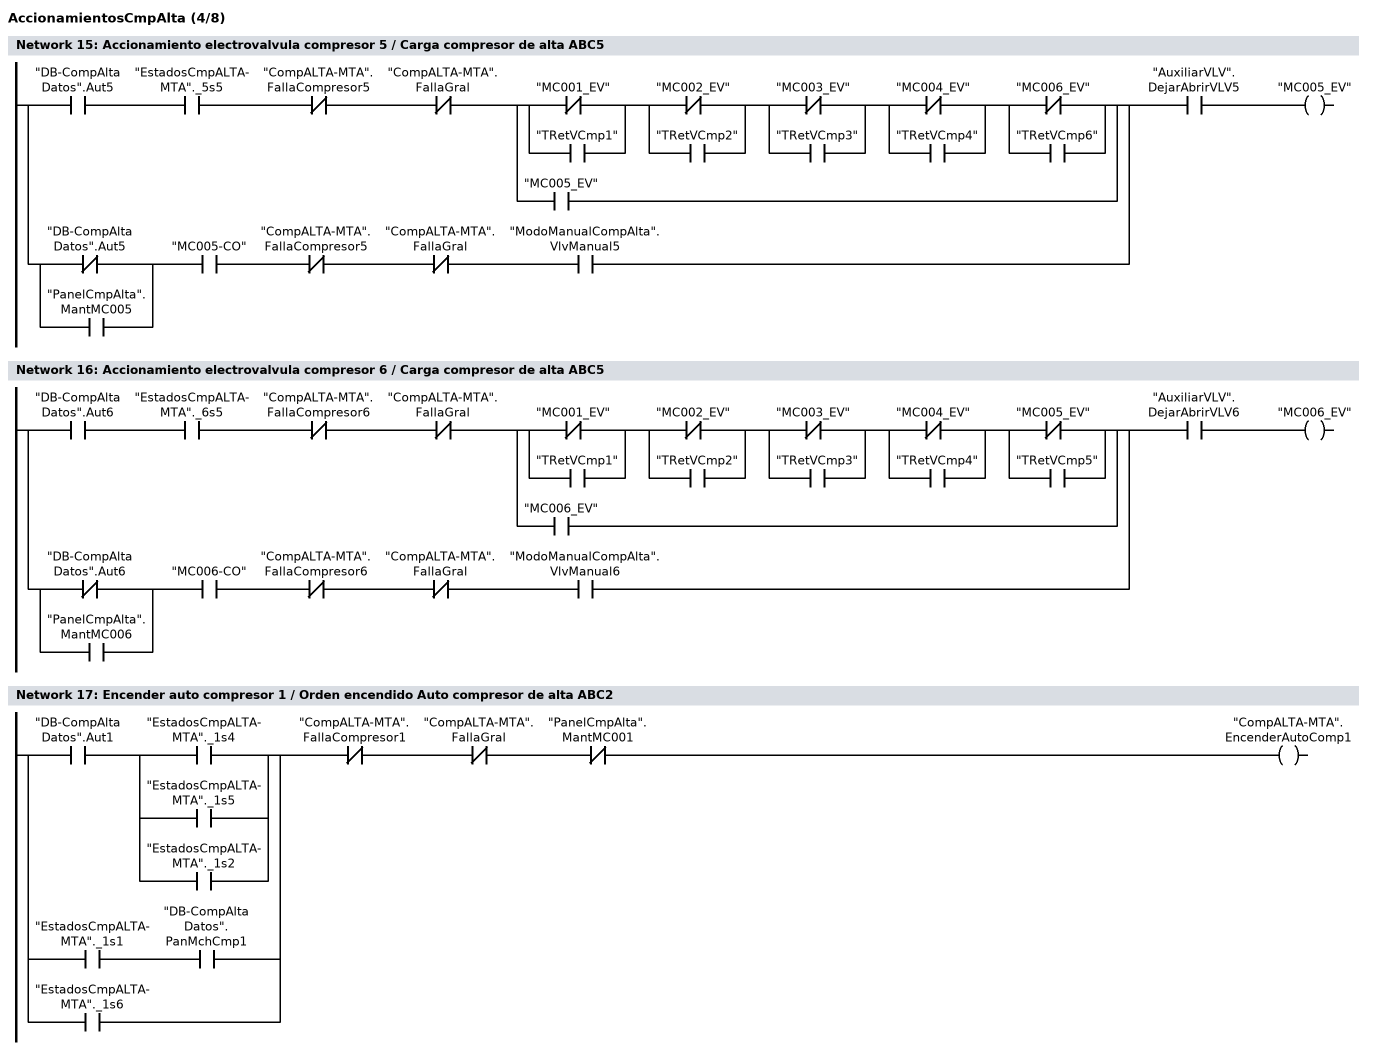
   RUNG wire#powerrail
      Contact( "DB-CompAltaDatos".Aut5 )
      Contact( "EstadosCmpALTA-MTA"._5s5 )
      I_Contact( "CompALTA-MTA".FallaCompresor5 )
      I_Contact( "CompALTA-MTA".FallaGral )
      wire#w1
      I_Contact( "MC001_EV" )
      wire#w2
      I_Contact( "MC002_EV" )
      wire#w3
      I_Contact( "MC003_EV" )
      wire#w4
      I_Contact( "MC004_EV" )
      wire#w5
      I_Contact( "MC006_EV" )
      wire#w6
      Contact( "AuxiliarVLV".DejarAbrirVLV5 )
      Coil( "MC005_EV" )
   END_RUNG
   RUNG wire#w1
      Contact( "TRetVCmp1" )
   END_RUNG wire#w2
   RUNG wire#w2
      Contact( "TRetVCmp2" )
   END_RUNG wire#w3
   RUNG wire#w3
      Contact( "TRetVCmp3" )
   END_RUNG wire#w4
   RUNG wire#w4
      Contact( "TRetVCmp4" )
   END_RUNG wire#w5
   RUNG wire#w5
      Contact( "TRetVCmp6" )
   END_RUNG wire#w6
   RUNG wire#w1
      Contact( "MC005_EV" )
   END_RUNG wire#w6
   RUNG wire#powerrail
      I_Contact( "DB-CompAltaDatos".Aut5 )
      wire#w7
      Contact( "MC005-CO" )
      I_Contact( "CompALTA-MTA".FallaCompresor5 )
      I_Contact( "CompALTA-MTA".FallaGral )
      Contact( "ModoManualCompAlta".VlvManual5 )
   END_RUNG wire#w6
   RUNG wire#powerrail
      Contact( "PanelCmpAlta".MantMC005 )
   END_RUNG wire#w7
   // the same network as SCL:
   "MC005_EV" := (("DB-CompAltaDatos".Aut5 AND "EstadosCmpALTA-MTA"._5s5 AND NOT "CompALTA-MTA".FallaCompresor5 AND NOT "CompALTA-MTA".FallaGral AND (((NOT "MC001_EV" OR "TRetVCmp1") AND (NOT "MC002_EV" OR "TRetVCmp2") AND (NOT "MC003_EV" OR "TRetVCmp3") AND (NOT "MC004_EV" OR "TRetVCmp4") AND (NOT "MC006_EV" OR "TRetVCmp6")) OR "MC005_EV")) OR ((NOT "DB-CompAltaDatos".Aut5 OR "PanelCmpAlta".MantMC005) AND "MC005-CO" AND NOT "CompALTA-MTA".FallaCompresor5 AND NOT "CompALTA-MTA".FallaGral AND "ModoManualCompAlta".VlvManual5)) AND "AuxiliarVLV".DejarAbrirVLV5;
END_REGION

REGION Network 16: Accionamiento electrovalvula compresor 6 / Carga compresor de alta ABC5
   RUNG wire#powerrail
      Contact( "DB-CompAltaDatos".Aut6 )
      Contact( "EstadosCmpALTA-MTA"._6s5 )
      I_Contact( "CompALTA-MTA".FallaCompresor6 )
      I_Contact( "CompALTA-MTA".FallaGral )
      wire#w1
      I_Contact( "MC001_EV" )
      wire#w2
      I_Contact( "MC002_EV" )
      wire#w3
      I_Contact( "MC003_EV" )
      wire#w4
      I_Contact( "MC004_EV" )
      wire#w5
      I_Contact( "MC005_EV" )
      wire#w6
      Contact( "AuxiliarVLV".DejarAbrirVLV6 )
      Coil( "MC006_EV" )
   END_RUNG
   RUNG wire#w1
      Contact( "TRetVCmp1" )
   END_RUNG wire#w2
   RUNG wire#w2
      Contact( "TRetVCmp2" )
   END_RUNG wire#w3
   RUNG wire#w3
      Contact( "TRetVCmp3" )
   END_RUNG wire#w4
   RUNG wire#w4
      Contact( "TRetVCmp4" )
   END_RUNG wire#w5
   RUNG wire#w5
      Contact( "TRetVCmp5" )
   END_RUNG wire#w6
   RUNG wire#w1
      Contact( "MC006_EV" )
   END_RUNG wire#w6
   RUNG wire#powerrail
      I_Contact( "DB-CompAltaDatos".Aut6 )
      wire#w7
      Contact( "MC006-CO" )
      I_Contact( "CompALTA-MTA".FallaCompresor6 )
      I_Contact( "CompALTA-MTA".FallaGral )
      Contact( "ModoManualCompAlta".VlvManual6 )
   END_RUNG wire#w6
   RUNG wire#powerrail
      Contact( "PanelCmpAlta".MantMC006 )
   END_RUNG wire#w7
   // the same network as SCL:
   "MC006_EV" := (("DB-CompAltaDatos".Aut6 AND "EstadosCmpALTA-MTA"._6s5 AND NOT "CompALTA-MTA".FallaCompresor6 AND NOT "CompALTA-MTA".FallaGral AND (((NOT "MC001_EV" OR "TRetVCmp1") AND (NOT "MC002_EV" OR "TRetVCmp2") AND (NOT "MC003_EV" OR "TRetVCmp3") AND (NOT "MC004_EV" OR "TRetVCmp4") AND (NOT "MC005_EV" OR "TRetVCmp5")) OR "MC006_EV")) OR ((NOT "DB-CompAltaDatos".Aut6 OR "PanelCmpAlta".MantMC006) AND "MC006-CO" AND NOT "CompALTA-MTA".FallaCompresor6 AND NOT "CompALTA-MTA".FallaGral AND "ModoManualCompAlta".VlvManual6)) AND "AuxiliarVLV".DejarAbrirVLV6;
END_REGION

REGION Network 17: Encender auto compresor 1 / Orden encendido Auto compresor de alta ABC2
   RUNG wire#powerrail
      Contact( "DB-CompAltaDatos".Aut1 )
      wire#w1
      Contact( "EstadosCmpALTA-MTA"._1s4 )
      wire#w2
      I_Contact( "CompALTA-MTA".FallaCompresor1 )
      I_Contact( "CompALTA-MTA".FallaGral )
      I_Contact( "PanelCmpAlta".MantMC001 )
      Coil( "CompALTA-MTA".EncenderAutoComp1 )
   END_RUNG
   RUNG wire#w1
      Contact( "EstadosCmpALTA-MTA"._1s5 )
   END_RUNG wire#w2
   RUNG wire#w1
      Contact( "EstadosCmpALTA-MTA"._1s2 )
   END_RUNG wire#w2
   RUNG wire#powerrail
      Contact( "EstadosCmpALTA-MTA"._1s1 )
      Contact( "DB-CompAltaDatos".PanMchCmp1 )
   END_RUNG wire#w2
   RUNG wire#powerrail
      Contact( "EstadosCmpALTA-MTA"._1s6 )
   END_RUNG wire#w2
   // the same network as SCL:
   "CompALTA-MTA".EncenderAutoComp1 := (("DB-CompAltaDatos".Aut1 AND ("EstadosCmpALTA-MTA"._1s4 OR "EstadosCmpALTA-MTA"._1s5 OR "EstadosCmpALTA-MTA"._1s2)) OR ("EstadosCmpALTA-MTA"._1s1 AND "DB-CompAltaDatos".PanMchCmp1) OR "EstadosCmpALTA-MTA"._1s6) AND NOT "CompALTA-MTA".FallaCompresor1 AND NOT "CompALTA-MTA".FallaGral AND NOT "PanelCmpAlta".MantMC001;
END_REGION

REGION Network 18: Encender auto compresor 2 / Orden encendido Auto compresor de alta ABC3
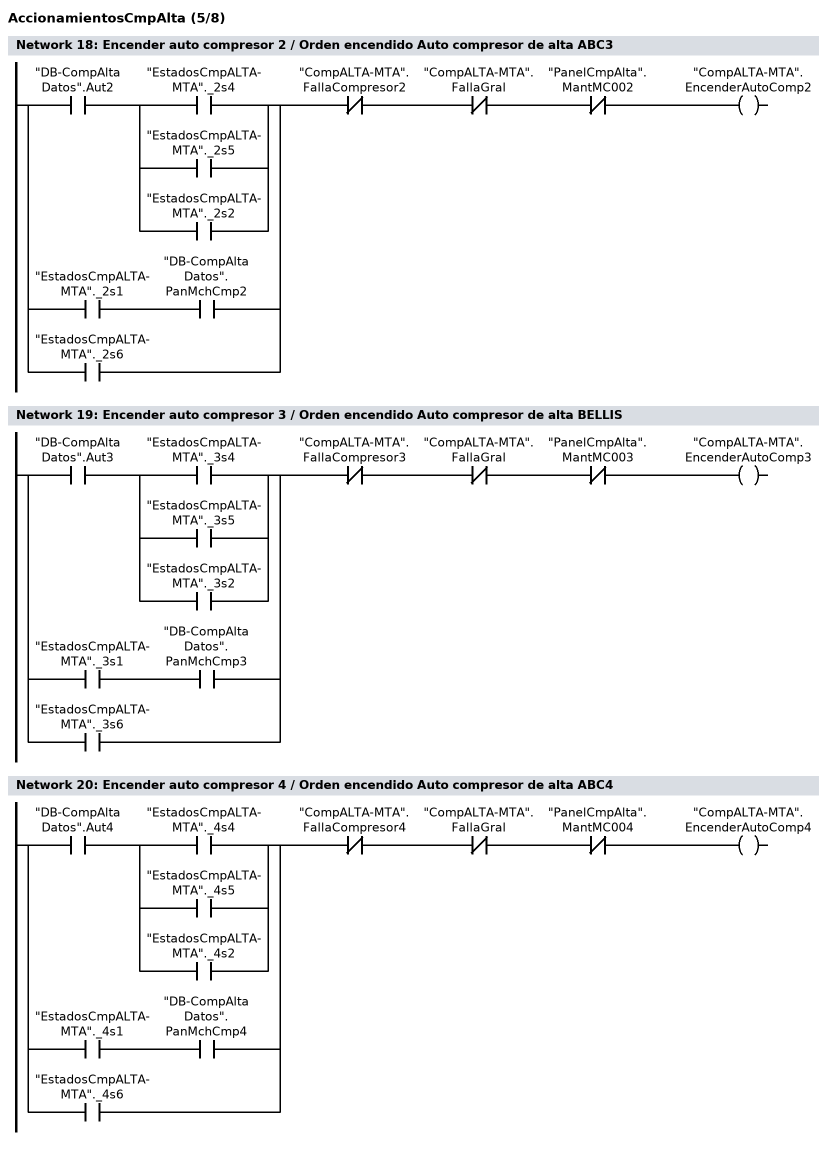
   RUNG wire#powerrail
      Contact( "DB-CompAltaDatos".Aut2 )
      wire#w1
      Contact( "EstadosCmpALTA-MTA"._2s4 )
      wire#w2
      I_Contact( "CompALTA-MTA".FallaCompresor2 )
      I_Contact( "CompALTA-MTA".FallaGral )
      I_Contact( "PanelCmpAlta".MantMC002 )
      Coil( "CompALTA-MTA".EncenderAutoComp2 )
   END_RUNG
   RUNG wire#w1
      Contact( "EstadosCmpALTA-MTA"._2s5 )
   END_RUNG wire#w2
   RUNG wire#w1
      Contact( "EstadosCmpALTA-MTA"._2s2 )
   END_RUNG wire#w2
   RUNG wire#powerrail
      Contact( "EstadosCmpALTA-MTA"._2s1 )
      Contact( "DB-CompAltaDatos".PanMchCmp2 )
   END_RUNG wire#w2
   RUNG wire#powerrail
      Contact( "EstadosCmpALTA-MTA"._2s6 )
   END_RUNG wire#w2
   // the same network as SCL:
   "CompALTA-MTA".EncenderAutoComp2 := (("DB-CompAltaDatos".Aut2 AND ("EstadosCmpALTA-MTA"._2s4 OR "EstadosCmpALTA-MTA"._2s5 OR "EstadosCmpALTA-MTA"._2s2)) OR ("EstadosCmpALTA-MTA"._2s1 AND "DB-CompAltaDatos".PanMchCmp2) OR "EstadosCmpALTA-MTA"._2s6) AND NOT "CompALTA-MTA".FallaCompresor2 AND NOT "CompALTA-MTA".FallaGral AND NOT "PanelCmpAlta".MantMC002;
END_REGION

REGION Network 19: Encender auto compresor 3 / Orden encendido Auto compresor de alta BELLIS
   RUNG wire#powerrail
      Contact( "DB-CompAltaDatos".Aut3 )
      wire#w1
      Contact( "EstadosCmpALTA-MTA"._3s4 )
      wire#w2
      I_Contact( "CompALTA-MTA".FallaCompresor3 )
      I_Contact( "CompALTA-MTA".FallaGral )
      I_Contact( "PanelCmpAlta".MantMC003 )
      Coil( "CompALTA-MTA".EncenderAutoComp3 )
   END_RUNG
   RUNG wire#w1
      Contact( "EstadosCmpALTA-MTA"._3s5 )
   END_RUNG wire#w2
   RUNG wire#w1
      Contact( "EstadosCmpALTA-MTA"._3s2 )
   END_RUNG wire#w2
   RUNG wire#powerrail
      Contact( "EstadosCmpALTA-MTA"._3s1 )
      Contact( "DB-CompAltaDatos".PanMchCmp3 )
   END_RUNG wire#w2
   RUNG wire#powerrail
      Contact( "EstadosCmpALTA-MTA"._3s6 )
   END_RUNG wire#w2
   // the same network as SCL:
   "CompALTA-MTA".EncenderAutoComp3 := (("DB-CompAltaDatos".Aut3 AND ("EstadosCmpALTA-MTA"._3s4 OR "EstadosCmpALTA-MTA"._3s5 OR "EstadosCmpALTA-MTA"._3s2)) OR ("EstadosCmpALTA-MTA"._3s1 AND "DB-CompAltaDatos".PanMchCmp3) OR "EstadosCmpALTA-MTA"._3s6) AND NOT "CompALTA-MTA".FallaCompresor3 AND NOT "CompALTA-MTA".FallaGral AND NOT "PanelCmpAlta".MantMC003;
END_REGION

REGION Network 20: Encender auto compresor 4 / Orden encendido Auto compresor de alta ABC4
   RUNG wire#powerrail
      Contact( "DB-CompAltaDatos".Aut4 )
      wire#w1
      Contact( "EstadosCmpALTA-MTA"._4s4 )
      wire#w2
      I_Contact( "CompALTA-MTA".FallaCompresor4 )
      I_Contact( "CompALTA-MTA".FallaGral )
      I_Contact( "PanelCmpAlta".MantMC004 )
      Coil( "CompALTA-MTA".EncenderAutoComp4 )
   END_RUNG
   RUNG wire#w1
      Contact( "EstadosCmpALTA-MTA"._4s5 )
   END_RUNG wire#w2
   RUNG wire#w1
      Contact( "EstadosCmpALTA-MTA"._4s2 )
   END_RUNG wire#w2
   RUNG wire#powerrail
      Contact( "EstadosCmpALTA-MTA"._4s1 )
      Contact( "DB-CompAltaDatos".PanMchCmp4 )
   END_RUNG wire#w2
   RUNG wire#powerrail
      Contact( "EstadosCmpALTA-MTA"._4s6 )
   END_RUNG wire#w2
   // the same network as SCL:
   "CompALTA-MTA".EncenderAutoComp4 := (("DB-CompAltaDatos".Aut4 AND ("EstadosCmpALTA-MTA"._4s4 OR "EstadosCmpALTA-MTA"._4s5 OR "EstadosCmpALTA-MTA"._4s2)) OR ("EstadosCmpALTA-MTA"._4s1 AND "DB-CompAltaDatos".PanMchCmp4) OR "EstadosCmpALTA-MTA"._4s6) AND NOT "CompALTA-MTA".FallaCompresor4 AND NOT "CompALTA-MTA".FallaGral AND NOT "PanelCmpAlta".MantMC004;
END_REGION

REGION Network 21: Encender auto compresor 5 / Orden encendido Auto compresor de alta ABC5
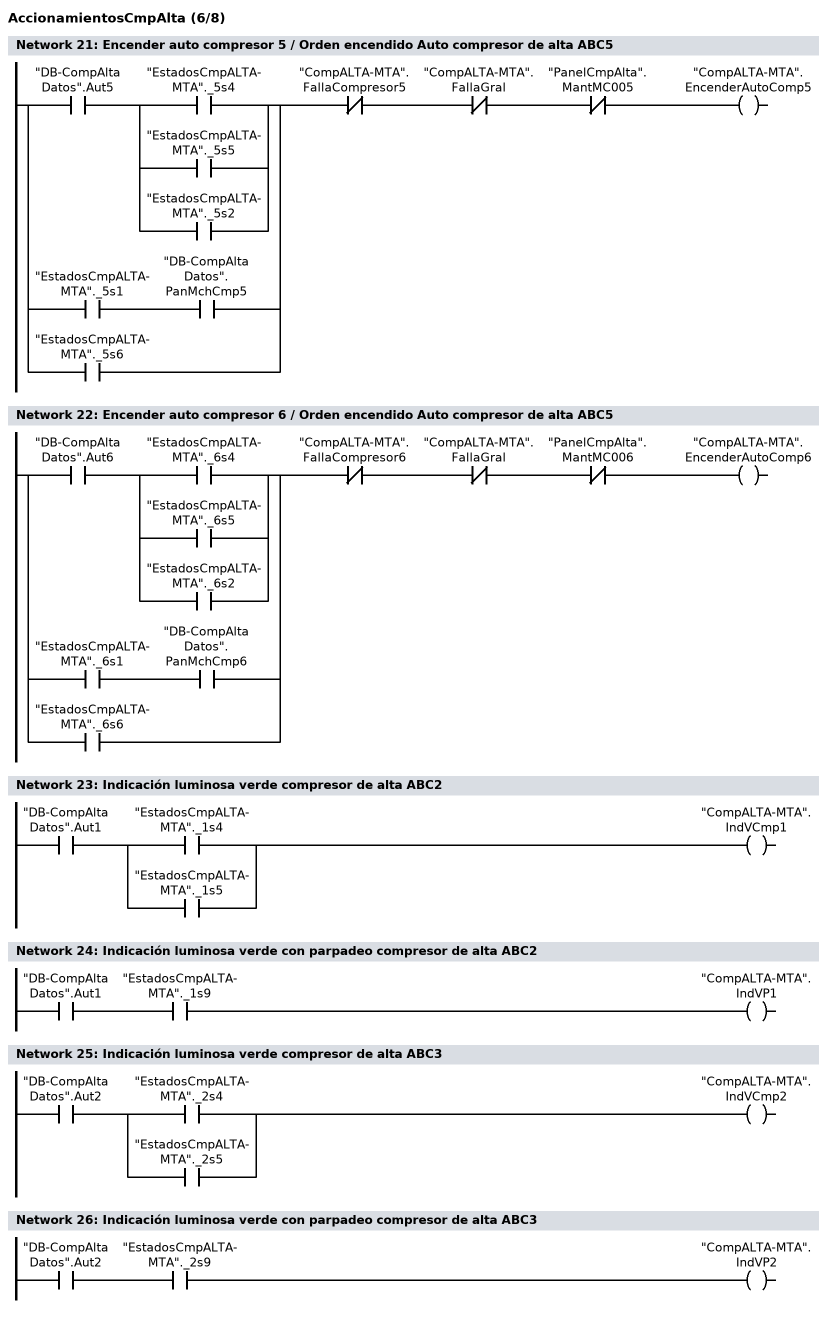
   RUNG wire#powerrail
      Contact( "DB-CompAltaDatos".Aut5 )
      wire#w1
      Contact( "EstadosCmpALTA-MTA"._5s4 )
      wire#w2
      I_Contact( "CompALTA-MTA".FallaCompresor5 )
      I_Contact( "CompALTA-MTA".FallaGral )
      I_Contact( "PanelCmpAlta".MantMC005 )
      Coil( "CompALTA-MTA".EncenderAutoComp5 )
   END_RUNG
   RUNG wire#w1
      Contact( "EstadosCmpALTA-MTA"._5s5 )
   END_RUNG wire#w2
   RUNG wire#w1
      Contact( "EstadosCmpALTA-MTA"._5s2 )
   END_RUNG wire#w2
   RUNG wire#powerrail
      Contact( "EstadosCmpALTA-MTA"._5s1 )
      Contact( "DB-CompAltaDatos".PanMchCmp5 )
   END_RUNG wire#w2
   RUNG wire#powerrail
      Contact( "EstadosCmpALTA-MTA"._5s6 )
   END_RUNG wire#w2
   // the same network as SCL:
   "CompALTA-MTA".EncenderAutoComp5 := (("DB-CompAltaDatos".Aut5 AND ("EstadosCmpALTA-MTA"._5s4 OR "EstadosCmpALTA-MTA"._5s5 OR "EstadosCmpALTA-MTA"._5s2)) OR ("EstadosCmpALTA-MTA"._5s1 AND "DB-CompAltaDatos".PanMchCmp5) OR "EstadosCmpALTA-MTA"._5s6) AND NOT "CompALTA-MTA".FallaCompresor5 AND NOT "CompALTA-MTA".FallaGral AND NOT "PanelCmpAlta".MantMC005;
END_REGION

REGION Network 22: Encender auto compresor 6 / Orden encendido Auto compresor de alta ABC5
   RUNG wire#powerrail
      Contact( "DB-CompAltaDatos".Aut6 )
      wire#w1
      Contact( "EstadosCmpALTA-MTA"._6s4 )
      wire#w2
      I_Contact( "CompALTA-MTA".FallaCompresor6 )
      I_Contact( "CompALTA-MTA".FallaGral )
      I_Contact( "PanelCmpAlta".MantMC006 )
      Coil( "CompALTA-MTA".EncenderAutoComp6 )
   END_RUNG
   RUNG wire#w1
      Contact( "EstadosCmpALTA-MTA"._6s5 )
   END_RUNG wire#w2
   RUNG wire#w1
      Contact( "EstadosCmpALTA-MTA"._6s2 )
   END_RUNG wire#w2
   RUNG wire#powerrail
      Contact( "EstadosCmpALTA-MTA"._6s1 )
      Contact( "DB-CompAltaDatos".PanMchCmp6 )
   END_RUNG wire#w2
   RUNG wire#powerrail
      Contact( "EstadosCmpALTA-MTA"._6s6 )
   END_RUNG wire#w2
   // the same network as SCL:
   "CompALTA-MTA".EncenderAutoComp6 := (("DB-CompAltaDatos".Aut6 AND ("EstadosCmpALTA-MTA"._6s4 OR "EstadosCmpALTA-MTA"._6s5 OR "EstadosCmpALTA-MTA"._6s2)) OR ("EstadosCmpALTA-MTA"._6s1 AND "DB-CompAltaDatos".PanMchCmp6) OR "EstadosCmpALTA-MTA"._6s6) AND NOT "CompALTA-MTA".FallaCompresor6 AND NOT "CompALTA-MTA".FallaGral AND NOT "PanelCmpAlta".MantMC006;
END_REGION

REGION Network 23: Indicación luminosa verde compresor de alta ABC2
   RUNG wire#powerrail
      Contact( "DB-CompAltaDatos".Aut1 )
      wire#w1
      Contact( "EstadosCmpALTA-MTA"._1s4 )
      wire#w2
      Coil( "CompALTA-MTA".IndVCmp1 )
   END_RUNG
   RUNG wire#w1
      Contact( "EstadosCmpALTA-MTA"._1s5 )
   END_RUNG wire#w2
   // the same network as SCL:
   "CompALTA-MTA".IndVCmp1 := "DB-CompAltaDatos".Aut1 AND ("EstadosCmpALTA-MTA"._1s4 OR "EstadosCmpALTA-MTA"._1s5);
END_REGION

REGION Network 24: Indicación luminosa verde con parpadeo compresor de alta ABC2
   RUNG wire#powerrail
      Contact( "DB-CompAltaDatos".Aut1 )
      Contact( "EstadosCmpALTA-MTA"._1s9 )
      Coil( "CompALTA-MTA".IndVP1 )
   END_RUNG
   // the same network as SCL:
   "CompALTA-MTA".IndVP1 := "DB-CompAltaDatos".Aut1 AND "EstadosCmpALTA-MTA"._1s9;
END_REGION

REGION Network 25: Indicación luminosa verde compresor de alta ABC3
   RUNG wire#powerrail
      Contact( "DB-CompAltaDatos".Aut2 )
      wire#w1
      Contact( "EstadosCmpALTA-MTA"._2s4 )
      wire#w2
      Coil( "CompALTA-MTA".IndVCmp2 )
   END_RUNG
   RUNG wire#w1
      Contact( "EstadosCmpALTA-MTA"._2s5 )
   END_RUNG wire#w2
   // the same network as SCL:
   "CompALTA-MTA".IndVCmp2 := "DB-CompAltaDatos".Aut2 AND ("EstadosCmpALTA-MTA"._2s4 OR "EstadosCmpALTA-MTA"._2s5);
END_REGION

REGION Network 26: Indicación luminosa verde con parpadeo compresor de alta ABC3
   RUNG wire#powerrail
      Contact( "DB-CompAltaDatos".Aut2 )
      Contact( "EstadosCmpALTA-MTA"._2s9 )
      Coil( "CompALTA-MTA".IndVP2 )
   END_RUNG
   // the same network as SCL:
   "CompALTA-MTA".IndVP2 := "DB-CompAltaDatos".Aut2 AND "EstadosCmpALTA-MTA"._2s9;
END_REGION

REGION Network 27: Indicación luminosa verde compresor de alta BELLIS
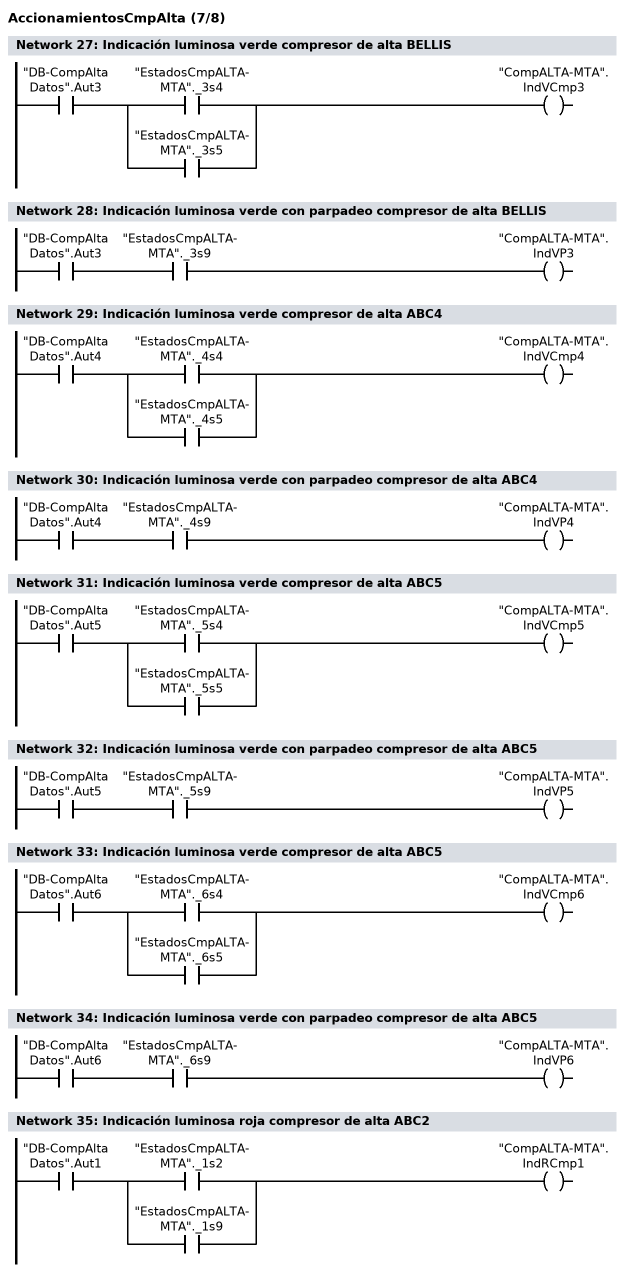
   RUNG wire#powerrail
      Contact( "DB-CompAltaDatos".Aut3 )
      wire#w1
      Contact( "EstadosCmpALTA-MTA"._3s4 )
      wire#w2
      Coil( "CompALTA-MTA".IndVCmp3 )
   END_RUNG
   RUNG wire#w1
      Contact( "EstadosCmpALTA-MTA"._3s5 )
   END_RUNG wire#w2
   // the same network as SCL:
   "CompALTA-MTA".IndVCmp3 := "DB-CompAltaDatos".Aut3 AND ("EstadosCmpALTA-MTA"._3s4 OR "EstadosCmpALTA-MTA"._3s5);
END_REGION

REGION Network 28: Indicación luminosa verde con parpadeo compresor de alta BELLIS
   RUNG wire#powerrail
      Contact( "DB-CompAltaDatos".Aut3 )
      Contact( "EstadosCmpALTA-MTA"._3s9 )
      Coil( "CompALTA-MTA".IndVP3 )
   END_RUNG
   // the same network as SCL:
   "CompALTA-MTA".IndVP3 := "DB-CompAltaDatos".Aut3 AND "EstadosCmpALTA-MTA"._3s9;
END_REGION

REGION Network 29: Indicación luminosa verde compresor de alta ABC4
   RUNG wire#powerrail
      Contact( "DB-CompAltaDatos".Aut4 )
      wire#w1
      Contact( "EstadosCmpALTA-MTA"._4s4 )
      wire#w2
      Coil( "CompALTA-MTA".IndVCmp4 )
   END_RUNG
   RUNG wire#w1
      Contact( "EstadosCmpALTA-MTA"._4s5 )
   END_RUNG wire#w2
   // the same network as SCL:
   "CompALTA-MTA".IndVCmp4 := "DB-CompAltaDatos".Aut4 AND ("EstadosCmpALTA-MTA"._4s4 OR "EstadosCmpALTA-MTA"._4s5);
END_REGION

REGION Network 30: Indicación luminosa verde con parpadeo compresor de alta ABC4
   RUNG wire#powerrail
      Contact( "DB-CompAltaDatos".Aut4 )
      Contact( "EstadosCmpALTA-MTA"._4s9 )
      Coil( "CompALTA-MTA".IndVP4 )
   END_RUNG
   // the same network as SCL:
   "CompALTA-MTA".IndVP4 := "DB-CompAltaDatos".Aut4 AND "EstadosCmpALTA-MTA"._4s9;
END_REGION

REGION Network 31: Indicación luminosa verde compresor de alta ABC5
   RUNG wire#powerrail
      Contact( "DB-CompAltaDatos".Aut5 )
      wire#w1
      Contact( "EstadosCmpALTA-MTA"._5s4 )
      wire#w2
      Coil( "CompALTA-MTA".IndVCmp5 )
   END_RUNG
   RUNG wire#w1
      Contact( "EstadosCmpALTA-MTA"._5s5 )
   END_RUNG wire#w2
   // the same network as SCL:
   "CompALTA-MTA".IndVCmp5 := "DB-CompAltaDatos".Aut5 AND ("EstadosCmpALTA-MTA"._5s4 OR "EstadosCmpALTA-MTA"._5s5);
END_REGION

REGION Network 32: Indicación luminosa verde con parpadeo compresor de alta ABC5
   RUNG wire#powerrail
      Contact( "DB-CompAltaDatos".Aut5 )
      Contact( "EstadosCmpALTA-MTA"._5s9 )
      Coil( "CompALTA-MTA".IndVP5 )
   END_RUNG
   // the same network as SCL:
   "CompALTA-MTA".IndVP5 := "DB-CompAltaDatos".Aut5 AND "EstadosCmpALTA-MTA"._5s9;
END_REGION

REGION Network 33: Indicación luminosa verde compresor de alta ABC5
   RUNG wire#powerrail
      Contact( "DB-CompAltaDatos".Aut6 )
      wire#w1
      Contact( "EstadosCmpALTA-MTA"._6s4 )
      wire#w2
      Coil( "CompALTA-MTA".IndVCmp6 )
   END_RUNG
   RUNG wire#w1
      Contact( "EstadosCmpALTA-MTA"._6s5 )
   END_RUNG wire#w2
   // the same network as SCL:
   "CompALTA-MTA".IndVCmp6 := "DB-CompAltaDatos".Aut6 AND ("EstadosCmpALTA-MTA"._6s4 OR "EstadosCmpALTA-MTA"._6s5);
END_REGION

REGION Network 34: Indicación luminosa verde con parpadeo compresor de alta ABC5
   RUNG wire#powerrail
      Contact( "DB-CompAltaDatos".Aut6 )
      Contact( "EstadosCmpALTA-MTA"._6s9 )
      Coil( "CompALTA-MTA".IndVP6 )
   END_RUNG
   // the same network as SCL:
   "CompALTA-MTA".IndVP6 := "DB-CompAltaDatos".Aut6 AND "EstadosCmpALTA-MTA"._6s9;
END_REGION

REGION Network 35: Indicación luminosa roja compresor de alta ABC2
   RUNG wire#powerrail
      Contact( "DB-CompAltaDatos".Aut1 )
      wire#w1
      Contact( "EstadosCmpALTA-MTA"._1s2 )
      wire#w2
      Coil( "CompALTA-MTA".IndRCmp1 )
   END_RUNG
   RUNG wire#w1
      Contact( "EstadosCmpALTA-MTA"._1s9 )
   END_RUNG wire#w2
   // the same network as SCL:
   "CompALTA-MTA".IndRCmp1 := "DB-CompAltaDatos".Aut1 AND ("EstadosCmpALTA-MTA"._1s2 OR "EstadosCmpALTA-MTA"._1s9);
END_REGION

REGION Network 36: Indicación luminosa roja compresor de alta ABC3
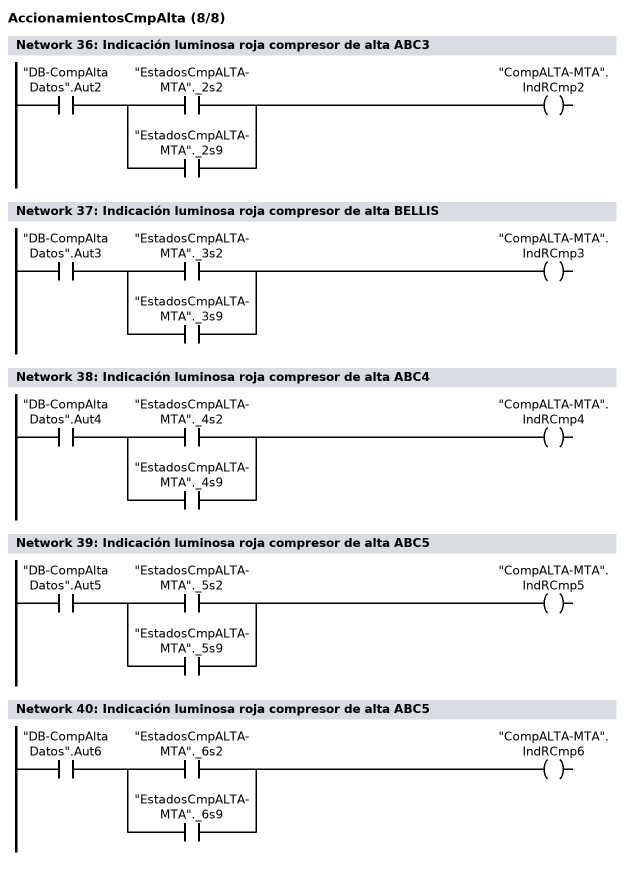
   RUNG wire#powerrail
      Contact( "DB-CompAltaDatos".Aut2 )
      wire#w1
      Contact( "EstadosCmpALTA-MTA"._2s2 )
      wire#w2
      Coil( "CompALTA-MTA".IndRCmp2 )
   END_RUNG
   RUNG wire#w1
      Contact( "EstadosCmpALTA-MTA"._2s9 )
   END_RUNG wire#w2
   // the same network as SCL:
   "CompALTA-MTA".IndRCmp2 := "DB-CompAltaDatos".Aut2 AND ("EstadosCmpALTA-MTA"._2s2 OR "EstadosCmpALTA-MTA"._2s9);
END_REGION

REGION Network 37: Indicación luminosa roja compresor de alta BELLIS
   RUNG wire#powerrail
      Contact( "DB-CompAltaDatos".Aut3 )
      wire#w1
      Contact( "EstadosCmpALTA-MTA"._3s2 )
      wire#w2
      Coil( "CompALTA-MTA".IndRCmp3 )
   END_RUNG
   RUNG wire#w1
      Contact( "EstadosCmpALTA-MTA"._3s9 )
   END_RUNG wire#w2
   // the same network as SCL:
   "CompALTA-MTA".IndRCmp3 := "DB-CompAltaDatos".Aut3 AND ("EstadosCmpALTA-MTA"._3s2 OR "EstadosCmpALTA-MTA"._3s9);
END_REGION

REGION Network 38: Indicación luminosa roja compresor de alta ABC4
   RUNG wire#powerrail
      Contact( "DB-CompAltaDatos".Aut4 )
      wire#w1
      Contact( "EstadosCmpALTA-MTA"._4s2 )
      wire#w2
      Coil( "CompALTA-MTA".IndRCmp4 )
   END_RUNG
   RUNG wire#w1
      Contact( "EstadosCmpALTA-MTA"._4s9 )
   END_RUNG wire#w2
   // the same network as SCL:
   "CompALTA-MTA".IndRCmp4 := "DB-CompAltaDatos".Aut4 AND ("EstadosCmpALTA-MTA"._4s2 OR "EstadosCmpALTA-MTA"._4s9);
END_REGION

REGION Network 39: Indicación luminosa roja compresor de alta ABC5
   RUNG wire#powerrail
      Contact( "DB-CompAltaDatos".Aut5 )
      wire#w1
      Contact( "EstadosCmpALTA-MTA"._5s2 )
      wire#w2
      Coil( "CompALTA-MTA".IndRCmp5 )
   END_RUNG
   RUNG wire#w1
      Contact( "EstadosCmpALTA-MTA"._5s9 )
   END_RUNG wire#w2
   // the same network as SCL:
   "CompALTA-MTA".IndRCmp5 := "DB-CompAltaDatos".Aut5 AND ("EstadosCmpALTA-MTA"._5s2 OR "EstadosCmpALTA-MTA"._5s9);
END_REGION

REGION Network 40: Indicación luminosa roja compresor de alta ABC5
   RUNG wire#powerrail
      Contact( "DB-CompAltaDatos".Aut6 )
      wire#w1
      Contact( "EstadosCmpALTA-MTA"._6s2 )
      wire#w2
      Coil( "CompALTA-MTA".IndRCmp6 )
   END_RUNG
   RUNG wire#w1
      Contact( "EstadosCmpALTA-MTA"._6s9 )
   END_RUNG wire#w2
   // the same network as SCL:
   "CompALTA-MTA".IndRCmp6 := "DB-CompAltaDatos".Aut6 AND ("EstadosCmpALTA-MTA"._6s2 OR "EstadosCmpALTA-MTA"._6s9);
END_REGION
END_FUNCTION

FUNCTION "PrioridadesReales" : Void   // FC41, LAD
{ S7_Optimized_Access := 'FALSE' }
VERSION : 0.1
BEGIN

REGION Network 1
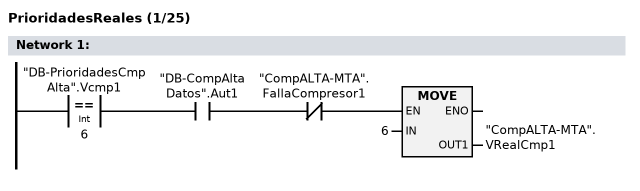
   RUNG wire#powerrail
      { S7_Templates := "SrcType := Int" } EQ_Contact(in1 := "DB-PrioridadesCmpAlta".Vcmp1, in2 := 6)
      Contact( "DB-CompAltaDatos".Aut1 )
      I_Contact( "CompALTA-MTA".FallaCompresor1 )
      { S7_GenerateENO := "TRUE" } Move(in := 6, out1 => "CompALTA-MTA".VRealCmp1)
   END_RUNG
   // the same network as SCL:
   IF ("DB-PrioridadesCmpAlta".Vcmp1 = 6) AND "DB-CompAltaDatos".Aut1 AND NOT "CompALTA-MTA".FallaCompresor1 THEN
       "CompALTA-MTA".VRealCmp1 := 6;
   END_IF;
END_REGION

REGION Network 2